// TIA Portal project "HEAT-1-CADIZ-V25" (V20) (continued)
VAR_GLOBAL   // PLC tag table "Robot Position"
   "tcpPosIniX_00" AT %I632.0 : Bool;   // $OUT[257]
   "tcpPosIniX_01" AT %I632.1 : Bool;
   "tcpPosIniX_02" AT %I632.2 : Bool;
   "tcpPosIniX_03" AT %I632.3 : Bool;
   "tcpPosIniX_04" AT %I632.4 : Bool;
   "tcpPosIniX_05" AT %I632.5 : Bool;
   "tcpPosIniX_06" AT %I632.6 : Bool;
   "tcpPosIniX_07" AT %I632.7 : Bool;
   "tcpPosIniX_08" AT %I633.0 : Bool;
   "tcpPosIniX_09" AT %I633.1 : Bool;
   "tcpPosIniX_10" AT %I633.2 : Bool;
   "tcpPosIniX_11" AT %I633.3 : Bool;
   "tcpPosIniX_12" AT %I633.4 : Bool;
   "tcpPosIniX_13" AT %I633.5 : Bool;
   "tcpPosIniX_14" AT %I633.6 : Bool;
   "tcpPosIniX_15" AT %I633.7 : Bool;
   "tcpPosIniX_16" AT %I634.0 : Bool;
   "tcpPosIniX_17" AT %I634.1 : Bool;
   "tcpPosIniX_18" AT %I634.2 : Bool;
   "tcpPosIniX_19" AT %I634.3 : Bool;
   "tcpPosIniX_20" AT %I634.4 : Bool;
   "tcpPosIniX_21" AT %I634.5 : Bool;
   "tcpPosIniX_22" AT %I634.6 : Bool;
   "tcpPosIniX_23" AT %I634.7 : Bool;
   "tcpPosIniX_24" AT %I635.0 : Bool;
   "tcpPosIniX_25" AT %I635.1 : Bool;
   "tcpPosIniX_26" AT %I635.2 : Bool;
   "tcpPosIniX_27" AT %I635.3 : Bool;
   "tcpPosIniX_28" AT %I635.4 : Bool;
   "tcpPosIniX_29" AT %I635.5 : Bool;
   "tcpPosIniX_30" AT %I635.6 : Bool;
   "tcpPosIniX_31" AT %I635.7 : Bool;
   "tcpPosIniY_00" AT %I636.0 : Bool;
   "tcpPosIniY_01" AT %I636.1 : Bool;
   "tcpPosIniY_02" AT %I636.2 : Bool;
   "tcpPosIniY_03" AT %I636.3 : Bool;
   "tcpPosIniY_04" AT %I636.4 : Bool;
   "tcpPosIniY_05" AT %I636.5 : Bool;
   "tcpPosIniY_06" AT %I636.6 : Bool;
   "tcpPosIniY_07" AT %I636.7 : Bool;
   "tcpPosIniY_08" AT %I637.0 : Bool;
   "tcpPosIniY_09" AT %I637.1 : Bool;
   "tcpPosIniY_10" AT %I637.2 : Bool;
   "tcpPosIniY_11" AT %I637.3 : Bool;
   "tcpPosIniY_12" AT %I637.4 : Bool;
   "tcpPosIniY_13" AT %I637.5 : Bool;
   "tcpPosIniY_14" AT %I637.6 : Bool;
   "tcpPosIniY_15" AT %I637.7 : Bool;
   "tcpPosIniY_16" AT %I638.0 : Bool;
   "tcpPosIniY_17" AT %I638.1 : Bool;
   "tcpPosIniY_18" AT %I638.2 : Bool;
   "tcpPosIniY_19" AT %I638.3 : Bool;
   "tcpPosIniY_20" AT %I638.4 : Bool;
   "tcpPosIniY_21" AT %I638.5 : Bool;
   "tcpPosIniY_22" AT %I638.6 : Bool;
   "tcpPosIniY_23" AT %I638.7 : Bool;
   "tcpPosIniY_24" AT %I639.0 : Bool;
   "tcpPosIniY_25" AT %I639.1 : Bool;
   "tcpPosIniY_26" AT %I639.2 : Bool;
   "tcpPosIniY_27" AT %I639.3 : Bool;
   "tcpPosIniY_28" AT %I639.4 : Bool;
   "tcpPosIniY_29" AT %I639.5 : Bool;
   "tcpPosIniY_30" AT %I639.6 : Bool;
   "tcpPosIniY_31" AT %I639.7 : Bool;
   "tcpPosIniZ_00" AT %I640.0 : Bool;
   "tcpPosIniZ_01" AT %I640.1 : Bool;
   "tcpPosIniZ_02" AT %I640.2 : Bool;
   "tcpPosIniZ_03" AT %I640.3 : Bool;
   "tcpPosIniZ_04" AT %I640.4 : Bool;
   "tcpPosIniZ_05" AT %I640.5 : Bool;
   "tcpPosIniZ_06" AT %I640.6 : Bool;
   "tcpPosIniZ_07" AT %I640.7 : Bool;
   "tcpPosIniZ_08" AT %I641.0 : Bool;
   "tcpPosIniZ_09" AT %I641.1 : Bool;
   "tcpPosIniZ_10" AT %I641.2 : Bool;
   "tcpPosIniZ_11" AT %I641.3 : Bool;
   "tcpPosIniZ_12" AT %I641.4 : Bool;
   "tcpPosIniZ_13" AT %I641.5 : Bool;
   "tcpPosIniZ_14" AT %I641.6 : Bool;
   "tcpPosIniZ_15" AT %I641.7 : Bool;
   "tcpPosIniZ_16" AT %I642.0 : Bool;
   "tcpPosIniZ_17" AT %I642.1 : Bool;
   "tcpPosIniZ_18" AT %I642.2 : Bool;
   "tcpPosIniZ_19" AT %I642.3 : Bool;
   "tcpPosIniZ_20" AT %I642.4 : Bool;
   "tcpPosIniZ_21" AT %I642.5 : Bool;
   "tcpPosIniZ_22" AT %I642.6 : Bool;
   "tcpPosIniZ_23" AT %I642.7 : Bool;
   "tcpPosIniZ_24" AT %I643.0 : Bool;
   "tcpPosIniZ_25" AT %I643.1 : Bool;
   "tcpPosIniZ_26" AT %I643.2 : Bool;
   "tcpPosIniZ_27" AT %I643.3 : Bool;
   "tcpPosIniZ_28" AT %I643.4 : Bool;
   "tcpPosIniZ_29" AT %I643.5 : Bool;
   "tcpPosIniZ_30" AT %I643.6 : Bool;
   "tcpPosIniZ_31" AT %I643.7 : Bool;
   "e1PosIni_00" AT %I644.0 : Bool;
   "e1PosIni_01" AT %I644.1 : Bool;
   "e1PosIni_02" AT %I644.2 : Bool;
   "e1PosIni_03" AT %I644.3 : Bool;
   "e1PosIni_04" AT %I644.4 : Bool;
   "e1PosIni_05" AT %I644.5 : Bool;
   "e1PosIni_06" AT %I644.6 : Bool;
   "e1PosIni_07" AT %I644.7 : Bool;
   "e1PosIni_08" AT %I645.0 : Bool;
   "e1PosIni_09" AT %I645.1 : Bool;
   "e1PosIni_10" AT %I645.2 : Bool;
   "e1PosIni_11" AT %I645.3 : Bool;
   "e1PosIni_12" AT %I645.4 : Bool;
   "e1PosIni_13" AT %I645.5 : Bool;
   "e1PosIni_14" AT %I645.6 : Bool;
   "e1PosIni_15" AT %I645.7 : Bool;
   "e1PosIni_16" AT %I646.0 : Bool;
   "e1PosIni_17" AT %I646.1 : Bool;
   "e1PosIni_18" AT %I646.2 : Bool;
   "e1PosIni_19" AT %I646.3 : Bool;
   "e1PosIni_20" AT %I646.4 : Bool;
   "e1PosIni_21" AT %I646.5 : Bool;
   "e1PosIni_22" AT %I646.6 : Bool;
   "e1PosIni_23" AT %I646.7 : Bool;
   "e1PosIni_24" AT %I647.0 : Bool;
   "e1PosIni_25" AT %I647.1 : Bool;
   "e1PosIni_26" AT %I647.2 : Bool;
   "e1PosIni_27" AT %I647.3 : Bool;
   "e1PosIni_28" AT %I647.4 : Bool;
   "e1PosIni_29" AT %I647.5 : Bool;
   "e1PosIni_30" AT %I647.6 : Bool;
   "e1PosIni_31" AT %I647.7 : Bool;
   "tcpPosFinX_00" AT %I648.0 : Bool;
   "tcpPosFinX_01" AT %I648.1 : Bool;
   "tcpPosFinX_02" AT %I648.2 : Bool;
   "tcpPosFinX_03" AT %I648.3 : Bool;
   "tcpPosFinX_04" AT %I648.4 : Bool;
   "tcpPosFinX_05" AT %I648.5 : Bool;
   "tcpPosFinX_06" AT %I648.6 : Bool;
   "tcpPosFinX_07" AT %I648.7 : Bool;
   "tcpPosFinX_08" AT %I649.0 : Bool;
   "tcpPosFinX_09" AT %I649.1 : Bool;
   "tcpPosFinX_10" AT %I649.2 : Bool;
   "tcpPosFinX_11" AT %I649.3 : Bool;
   "tcpPosFinX_12" AT %I649.4 : Bool;
   "tcpPosFinX_13" AT %I649.5 : Bool;
   "tcpPosFinX_14" AT %I649.6 : Bool;
   "tcpPosFinX_15" AT %I649.7 : Bool;
   "tcpPosFinX_16" AT %I650.0 : Bool;
   "tcpPosFinX_17" AT %I650.1 : Bool;
   "tcpPosFinX_18" AT %I650.2 : Bool;
   "tcpPosFinX_19" AT %I650.3 : Bool;
   "tcpPosFinX_20" AT %I650.4 : Bool;
   "tcpPosFinX_21" AT %I650.5 : Bool;
   "tcpPosFinX_22" AT %I650.6 : Bool;
   "tcpPosFinX_23" AT %I650.7 : Bool;
   "tcpPosFinX_24" AT %I651.0 : Bool;
   "tcpPosFinX_25" AT %I651.1 : Bool;
   "tcpPosFinX_26" AT %I651.2 : Bool;
   "tcpPosFinX_27" AT %I651.3 : Bool;
   "tcpPosFinX_28" AT %I651.4 : Bool;
   "tcpPosFinX_29" AT %I651.5 : Bool;
   "tcpPosFinX_30" AT %I651.6 : Bool;
   "tcpPosFinX_31" AT %I651.7 : Bool;
   "tcpPosFinY_00" AT %I652.0 : Bool;
   "tcpPosFinY_01" AT %I652.1 : Bool;
   "tcpPosFinY_02" AT %I652.2 : Bool;
   "tcpPosFinY_03" AT %I652.3 : Bool;
   "tcpPosFinY_04" AT %I652.4 : Bool;
   "tcpPosFinY_05" AT %I652.5 : Bool;
   "tcpPosFinY_06" AT %I652.6 : Bool;
   "tcpPosFinY_07" AT %I652.7 : Bool;
   "tcpPosFinY_08" AT %I653.0 : Bool;
   "tcpPosFinY_09" AT %I653.1 : Bool;
   "tcpPosFinY_10" AT %I653.2 : Bool;
   "tcpPosFinY_11" AT %I653.3 : Bool;
   "tcpPosFinY_12" AT %I653.4 : Bool;
   "tcpPosFinY_13" AT %I653.5 : Bool;
   "tcpPosFinY_14" AT %I653.6 : Bool;
   "tcpPosFinY_15" AT %I653.7 : Bool;
   "tcpPosFinY_16" AT %I654.0 : Bool;
   "tcpPosFinY_17" AT %I654.1 : Bool;
   "tcpPosFinY_18" AT %I654.2 : Bool;
   "tcpPosFinY_19" AT %I654.3 : Bool;
   "tcpPosFinY_20" AT %I654.4 : Bool;
   "tcpPosFinY_21" AT %I654.5 : Bool;
   "tcpPosFinY_22" AT %I654.6 : Bool;
   "tcpPosFinY_23" AT %I654.7 : Bool;
   "tcpPosFinY_24" AT %I655.0 : Bool;
   "tcpPosFinY_25" AT %I655.1 : Bool;
   "tcpPosFinY_26" AT %I655.2 : Bool;
   "tcpPosFinY_27" AT %I655.3 : Bool;
   "tcpPosFinY_28" AT %I655.4 : Bool;
   "tcpPosFinY_29" AT %I655.5 : Bool;
   "tcpPosFinY_30" AT %I655.6 : Bool;
   "tcpPosFinY_31" AT %I655.7 : Bool;
   "tcpPosE1_01" AT %I628.0 : Bool;
   "tcpPosE1_02" AT %I628.1 : Bool;
   "tcpPosE1_03" AT %I628.2 : Bool;
   "tcpPosE1_04" AT %I628.3 : Bool;
   "tcpPosE1_05" AT %I628.4 : Bool;
   "tcpPosE1_06" AT %I628.5 : Bool;
   "tcpPosE1_07" AT %I628.6 : Bool;
   "tcpPosE1_08" AT %I628.7 : Bool;
   "tcpPosE1_09" AT %I629.0 : Bool;
   "tcpPosE1_10" AT %I629.1 : Bool;
   "tcpPosE1_11" AT %I629.2 : Bool;
   "tcpPosE1_12" AT %I629.3 : Bool;
   "tcpPosE1_13" AT %I629.4 : Bool;
   "tcpPosE1_14" AT %I629.5 : Bool;
   "tcpPosE1_15" AT %I629.6 : Bool;
   "tcpPosE1_16" AT %I629.7 : Bool;
   "tcpPosE1_17" AT %I630.0 : Bool;
   "tcpPosE1_18" AT %I630.1 : Bool;
   "tcpPosE1_19" AT %I630.2 : Bool;
   "tcpPosE1_20" AT %I630.3 : Bool;
   "tcpPosE1_21" AT %I630.4 : Bool;
   "tcpPosE1_22" AT %I630.5 : Bool;
   "tcpPosE1_23" AT %I630.6 : Bool;
   "tcpPosE1_24" AT %I630.7 : Bool;
   "tcpPosE1_25" AT %I631.0 : Bool;
   "tcpPosE1_26" AT %I631.1 : Bool;
   "tcpPosE1_27" AT %I631.2 : Bool;
   "tcpPosE1_28" AT %I631.3 : Bool;
   "tcpPosE1_29" AT %I631.4 : Bool;
   "tcpPosE1_30" AT %I631.5 : Bool;
   "tcpPosE1_31" AT %I631.6 : Bool;
   "tcpPosE1_32" AT %I631.7 : Bool;
   "tcpPosIniX_rawLe32" AT %ID632 : DWord;
   "tcpPosIniY_rawLe32" AT %ID636 : DWord;
   "tcpPosIniZ_rawLe32" AT %ID640 : DWord;
   "tcpPosFinX_rawLe32" AT %ID648 : DWord;
   "tcpPosFinY_rawLe32" AT %ID652 : DWord;
   "e1_rawLe32" AT %ID628 : DWord;
   "e1PosIni_rawLe32" AT %ID644 : DWord;
   "tcpPosFinZ_rawLe32" AT %ID656 : DWord;
   "e1PosFin_rawLe32" AT %ID660 : DWord;
END_VAR

VAR_GLOBAL   // PLC tag table "Tool Change"
   "dockSensorToolYugoInPosition" AT %I150.0 : Bool;   // DETECTOR_YUGO_LP
   "dockSensorCoverYugoClosed" AT %I150.1 : Bool;   // TAPA_CERRADA_YUGO_LP
   "dockSensorCoverOpen" AT %I160.0 : Bool;   // TAPA_ABIERTA_YUGO_LP
   "dockValveV2UnlockOnYugo" AT %Q171.2 : Bool;   // SOLTAR_HERRAMIENTA_YUGO_LP / CAMBIA A FALSE
   "dockValveCoverOpenOn" AT %Q170.0 : Bool;   // ABRIR_TAPA_YUGO_LP
   "dockValveCoverCloseOn" AT %Q170.1 : Bool;   // CERRAR_TAPA_YUGO_LP
   "robotSensorMpsUnlocked" AT %I200.0 : Bool;   // INTERCAMBIO_DESBLOQUEADO_LR
   "robotSensorMpsLocked" AT %I200.1 : Bool;   // INTERCAMBIO_BLOQUEADO_LR
   "robotSensorMpsCoupled" AT %I200.2 : Bool;   // HERRAMIENTA_PUESTA_LR /AL COLOCAR METAL
   "robotSensorMpsCtrlAirPressureOk" AT %I200.3 : Bool;   // PRESION_CORRECTA_LR
   "toolReqId_01" AT %Q618.1 : Bool;   // INKUKA_DETECTOR_HERRAMIENTA
   "toolReqId_02" AT %Q618.2 : Bool;   // INKUKA_TAPA_CERRADA_YUGO
   "toolReqId_03" AT %Q618.3 : Bool;   // INKUKA_TAPA_ABIERTA_YUGO
   "toolReqId_04" AT %Q618.4 : Bool;   // INKUKA_INTERCAMBIO_DESBLOQUEADO
   "toolReqId_05" AT %Q618.5 : Bool;   // INKUKA_INTERCAMBIO_BLOQUEADO
   "toolReqId_06" AT %Q618.6 : Bool;   // INKUKA_HERRAMIENTA_PUESTA /AL COLOCAR util met
   "toolReqId_07" AT %Q618.7 : Bool;
   "kukaCmdUnlockMpsYugo" AT %I696.0 : Bool;   // OUTKUKA_SOLTAR_HERRAMIENTA_YUGO
   "kukaCmdOpenCover" AT %I696.1 : Bool;   // OUTKUKA_ABRIR_TAPA_YUGO
   "kukaCmdCloseCover" AT %I696.2 : Bool;   // OUTKUKA_CERRAR_TAPA_YUGO
   "V1_B14_S2" AT %Q0.0 : Bool;   // Anticolision - OPR
   "V1_B12_S4" AT %Q0.1 : Bool;   // Mps Bloqueo SIL 2
   "V2_B14_S2" AT %Q0.2 : Bool;
   "V2_B12_S4" AT %Q0.3 : Bool;
   "toolReqId_00" AT %Q618.0 : Bool;
   "toolReqId_08" AT %Q619.0 : Bool;
   "toolReqId_09" AT %Q619.1 : Bool;
   "toolReqId_10" AT %Q619.2 : Bool;
   "toolReqId_11" AT %Q619.3 : Bool;
   "toolReqId_12" AT %Q619.4 : Bool;
   "toolReqId_13" AT %Q619.5 : Bool;
   "toolReqId_14" AT %Q619.6 : Bool;
   "toolReqId_15" AT %Q619.7 : Bool;
   "toolReqId" AT %QW618 : Word;
   "baseReqId" AT %QW620 : Word;
   "kukaFeedbackDockToolYugoInPosition" AT %Q696.4 : Bool;   // $IN[773]
   "kukaFeedbackDockYugoCoverClosed" AT %Q696.5 : Bool;
   "kukaFeedbackDockYugoCoverOpen" AT %Q696.6 : Bool;
   "kukaFeedbackRobotMpsUnlocked" AT %Q696.0 : Bool;   // $IN[769]
   "kukaFeedbackRobotMpsLocked" AT %Q696.1 : Bool;
   "kukaFeedbackRobotMpsCoupled" AT %Q696.2 : Bool;
   "kukaFeedbackRobotMpsCtrlAirPressureOk" AT %Q696.3 : Bool;
   "dockValveV2UnlockOnPepa" AT %Q171.4 : Bool;   // SOLTAR_HERRAMIENTA_PEPA
   "dockSensorToolPepaInPosition" AT %I150.2 : Bool;
   "kukaCmdSafeForChange" AT %I696.3 : Bool;   // $OUT[772]
   "kukaCmdUnlockMpsPepa" AT %I696.4 : Bool;   // $OUT[773]
   "kukaCmdOpenCoverPepa" AT %I696.5 : Bool;   // $OUT[774]
   "kukaCmdUnlockMpsMarker" AT %I696.7 : Bool;   // $OUT[775]
   "kukaCmdOpenCoverMarker" AT %I697.0 : Bool;   // $OUT[776]
   "kukaCmdCloseCoverMarker" AT %I697.1 : Bool;   // $OUT[777]
   "kukaCmdUnlockMpsGocator" AT %I697.2 : Bool;
   "kukaCmdOpenCoverGocator" AT %I697.3 : Bool;
   "kukaCmdCloseCoverGocator" AT %I697.4 : Bool;
   "kukaCmdCloseCoverPepa" AT %I696.6 : Bool;
   "kukaCmdUnlockMpsPole" AT %I697.5 : Bool;
   "kukaCmdOpenCoverPole" AT %I697.6 : Bool;
   "kukaCmdCloseCoverPole" AT %I697.7 : Bool;
   "kukaFeedbackDockToolPepaInPosition" AT %Q696.7 : Bool;
   "kukaFeedbackDockPepaCoverClosed" AT %Q697.0 : Bool;
   "kukaFeedbackDockPepaCoverOpen" AT %Q697.1 : Bool;
   "kukaFeedbackDockToolMarkerInPosition" AT %Q697.2 : Bool;
   "kukaFeedbackDockMarkerCoverClosed" AT %Q697.3 : Bool;
   "kukaFeedbackDockMarkerCoverOpen" AT %Q697.4 : Bool;
   "kukaFeedbackDockToolGocatorInPosition" AT %Q697.5 : Bool;
   "kukaFeedbackDockGocatorCoverClosed" AT %Q697.6 : Bool;
   "kukaFeedbackDockGocatorCoverOpen" AT %Q697.7 : Bool;
   "kukaFeedbackDockToolPoleInPosition" AT %Q698.0 : Bool;
   "kukaFeedbackDockPoleCoverClosed" AT %Q698.1 : Bool;
   "kukaFeedbackDockPoleCoverOpen" AT %Q698.2 : Bool;
   "dockSensorCoverPepaClosed" AT %I150.3 : Bool;
   "dockSensorToolPoleInPosition" AT %I150.4 : Bool;
   "dockSensorToolMarkerInPosition" AT %I150.6 : Bool;
   "dockSensorToolGocatorInPosition" AT %I151.0 : Bool;
   "pruebaHerramienta2enStand" AT %I151.2 : Bool;
   "pruebaHerramienta1enStand" AT %I151.1 : Bool;
   "pruebaHerramienta3enStand" AT %I151.3 : Bool;
   "pruebaHerramienta4enStand" AT %I151.4 : Bool;
   "pruebaHerramient54enStand" AT %I150.7 : Bool;
   "dockSensorTooPole%I150.5InPosition" AT %I150.5 : Bool;
END_VAR

VAR_GLOBAL   // PLC tag table "General"
   "ALM_PRESS_SENSOR" AT %I10.0 : Bool;   // Pressure-sensor alarm
   "CMD_TANK_FILL" AT %Q30.0 : Bool;   // LLENAR CUBA
   "CMD_TANK_DRAIN" AT %Q30.1 : Bool;   // VACIAR CUBA
   "RECIRCULACION" AT %Q30.2 : Bool;   // CONMUTADOR MANUAL / cambiado a recirculacion
END_VAR

VAR_GLOBAL   // PLC tag table "Tag table_1"
   "Sensor_plato_giro_1" AT %I410.0 : Bool;
   "Sensor_Plato_giro_2" AT %I410.1 : Bool;
   "Sensor_plato_giro_3" AT %I410.2 : Bool;
   "Sensor_ADN_bastidor_bloqueado_1" AT %I410.3 : Bool;
   "Sensor_ADN_bastidor_desbloqueado_1" AT %I410.4 : Bool;
   "Sensor_ADN_bastidor_bloqueado_2" AT %I410.5 : Bool;
   "Sensor_ADN_bastidor_desbloqueado_2" AT %I410.6 : Bool;
   "SENSOR_CRDSNU_BASTIDOR_BLOQUEADO_1" AT %I410.7 : Bool;
   "SENSOR_CRDSNU_BASTIDOR_DESBLOQUEADO_1" AT %I411.0 : Bool;
   "SENSOR_CRDSNU_BASTIDOR_BLOQUEADO_2" AT %I411.1 : Bool;
   "SENSOR_CRDSNU_BASTIDOR_DESBLOQUEADO_2" AT %I411.2 : Bool;
   "SENSOR_DSBG_BASTIDOR_ARRIBA_1" AT %I411.3 : Bool;
   "SENSOR_DSBG_BASTIDOR_ABAJO_1" AT %I411.4 : Bool;
   "SENSOR_DSBG_BASTIDOR_ARRIBA_2" AT %I411.5 : Bool;
   "SENSOR_DSBG_BASTIDOR_ABAJO_2" AT %I411.6 : Bool;
   "PULSADOR_SUBIR_1" AT %I412.0 : Bool;
   "PULSADOR_BAJAR_1" AT %I412.1 : Bool;
   "PULSADOR_SUBIR_2" AT %I412.2 : Bool;
   "PULSADOR_BAJAR_2" AT %I412.3 : Bool;
   "VALVULA_52_BIESTABLE_11" AT %Q420.0 : Bool;
   "VALVULA_52_BIESTABLE_12" AT %Q420.1 : Bool;
   "VALVULA_52_BIESTABLE_21" AT %Q420.2 : Bool;
   "VALVULA_52_BIESTABLE_22" AT %Q420.3 : Bool;
   "VÁLVULA_52_MONOESTABLE_1" AT %Q420.4 : Bool;
   "VÁLVULA_52_MONOESTABLE_2" AT %Q420.5 : Bool;
   "VÁLVULA_52_MONOESTABLE_3" AT %Q420.6 : Bool;
   "VÁLVULA_52_MONOESTABLE_4" AT %Q420.7 : Bool;
   "VÁLVULA_52_MONOESTABLE_5" AT %Q421.0 : Bool;
   "SENSOR_DSBG_BASTIDOR_ABAJO_3" AT %I411.7 : Bool;
   "PULSADOR_BAJAR_3" AT %I412.4 : Bool;
   "PULSADOR_BAJAR_4" AT %I412.5 : Bool;
   "PULSADOR_BAJAR_5" AT %I412.6 : Bool;
   "PULSADOR_BAJAR_6" AT %I412.7 : Bool;
   "PULSADOR_BAJAR_7" AT %I413.0 : Bool;
   "PULSADOR_BAJAR_8" AT %I413.1 : Bool;
   "PULSADOR_BAJAR_9" AT %I413.2 : Bool;
   "PULSADOR_BAJAR_10" AT %I413.3 : Bool;
   "PULSADOR_BAJAR_11" AT %I413.4 : Bool;
   "PULSADOR_BAJAR_12" AT %I413.5 : Bool;
   "PULSADOR_BAJAR_13" AT %I413.6 : Bool;
   "PULSADOR_BAJAR_14" AT %I413.7 : Bool;
   "VÁLVULA_52_MONOESTABLE_6" AT %Q421.1 : Bool;
   "VÁLVULA_52_MONOESTABLE_7" AT %Q421.2 : Bool;
   "VÁLVULA_52_MONOESTABLE_8" AT %Q421.3 : Bool;
   "VÁLVULA_52_MONOESTABLE_9" AT %Q421.4 : Bool;
   "VÁLVULA_52_MONOESTABLE_10" AT %Q421.5 : Bool;
   "VÁLVULA_52_MONOESTABLE_11" AT %Q421.6 : Bool;
   "VÁLVULA_52_MONOESTABLE_12" AT %Q421.7 : Bool;
   "VÁLVULA_52_MONOESTABLE_13" AT %Q422.0 : Bool;
   "VÁLVULA_52_MONOESTABLE_14" AT %Q422.1 : Bool;
   "VÁLVULA_52_MONOESTABLE_15" AT %Q422.2 : Bool;
   "VÁLVULA_52_MONOESTABLE_16" AT %Q422.3 : Bool;
   "VÁLVULA_52_MONOESTABLE_17" AT %Q422.4 : Bool;
   "VÁLVULA_52_MONOESTABLE_18" AT %Q422.5 : Bool;
   "VÁLVULA_52_MONOESTABLE_19" AT %Q422.6 : Bool;
   "VÁLVULA_52_MONOESTABLE_20" AT %Q422.7 : Bool;
   "VÁLVULA_52_MONOESTABLE_21" AT %Q423.0 : Bool;
   "VÁLVULA_52_MONOESTABLE_22" AT %Q423.1 : Bool;
   "VÁLVULA_52_MONOESTABLE_23" AT %Q423.2 : Bool;
   "VÁLVULA_52_MONOESTABLE_24" AT %Q423.3 : Bool;
   "VÁLVULA_52_MONOESTABLE_25" AT %Q423.4 : Bool;
   "VÁLVULA_52_MONOESTABLE_26" AT %Q423.5 : Bool;
   "VÁLVULA_52_MONOESTABLE_27" AT %Q423.6 : Bool;
   "VÁLVULA_52_MONOESTABLE_28" AT %Q423.7 : Bool;
END_VAR

TYPE "UDT_Dock"
   STRUCT
      Sensor : Struct
         CoverOpen : Bool;
         CoverClosed : Bool;
         ToolInPosition : Bool;
      END_STRUCT;
      Valve : Struct
         CoverOpenOn : Bool;
         CoverCloseOn : Bool;
         V2UnlockOn : Bool;
      END_STRUCT;
   END_STRUCT;
END_TYPE

TYPE "UDT_RobotMps"
   STRUCT
      Sensor : Struct
         Coupled : Bool;
         Locked : Bool;
         Unlocked : Bool;
         CtrlAirPressureOk : Bool;
      END_STRUCT;
   END_STRUCT;
END_TYPE

// folder: 10. System

DATA_BLOCK "HMI_CUBA_DB"   // DB17
{ S7_Optimized_Access := 'TRUE' }
VERSION : 0.1
// stored: InstanceOfName HMI_CUBA
"HMI_CUBA"
BEGIN
END_DATA_BLOCK

DATA_BLOCK "instKukaControlSeq_DB"   // DB20
{ S7_Optimized_Access := 'TRUE' }
VERSION : 0.1
// stored: InstanceOfName KukaControlSeq
"KukaControlSeq"
BEGIN
END_DATA_BLOCK

DATA_BLOCK "GIRO_POSITIVO_DB"   // DB27
{ S7_Optimized_Access := 'TRUE' }
VERSION : 0.1
// stored: InstanceOfName GIRO_POSITIVO
"GIRO_POSITIVO"
BEGIN
END_DATA_BLOCK

DATA_BLOCK "GIRO_NEGATIVO_1_DB"   // DB28
{ S7_Optimized_Access := 'TRUE' }
VERSION : 0.1
// stored: InstanceOfName GIRO_NEGATIVO_1
"GIRO_NEGATIVO_1"
BEGIN
END_DATA_BLOCK

// folder: 10. System/DbsInstancia

DATA_BLOCK "InstKukaControlSeq"   // DB14
{ S7_Optimized_Access := 'TRUE' }
VERSION : 0.1
// stored: InstanceOfName KukaControlSeq
"KukaControlSeq"
BEGIN
END_DATA_BLOCK

DATA_BLOCK "InstSupervisorSeq"   // DB15
{ S7_Optimized_Access := 'TRUE' }
VERSION : 0.1
// stored: InstanceOfName SupervisorSeq
"SupervisorSeq"
BEGIN
END_DATA_BLOCK

DATA_BLOCK "InstSeqManager"   // DB16
{ S7_Optimized_Access := 'TRUE' }
VERSION : 0.1
// stored: InstanceOfName SeqManager
"SeqManager"
BEGIN
END_DATA_BLOCK

DATA_BLOCK "AutoExtSeq_DB"   // DB18
{ S7_Optimized_Access := 'TRUE' }
VERSION : 0.1
// stored: InstanceOfName AutoExtSeq
"AutoExtSeq"
BEGIN
END_DATA_BLOCK

DATA_BLOCK "instSupervisorSeq_DB"   // DB21
{ S7_Optimized_Access := 'TRUE' }
VERSION : 0.1
// stored: InstanceOfName SupervisorSeq
"SupervisorSeq"
BEGIN
END_DATA_BLOCK

// folder: 10. System/DbsOpcUa

DATA_BLOCK "PlcStatus"   // DB4
{ S7_Optimized_Access := 'TRUE' }
VERSION : 0.1
   VAR
      "- FOR  KUKACONTROL-" : Bool;
      mode : Struct
         effective : UInt;
         ready : Bool;
      END_STRUCT;
      active : Struct
         baseId : UInt;
         toolId : UInt;
         profileId : UInt;
      END_STRUCT;
      exec : Struct
         ackSeq : UInt;
         accepted : Bool;
         busy : Bool;
         done : Bool;
         error : Bool;
         errorCode : UDInt;
         cancelAck : Bool;
         pauseAck : Bool;
         resumeAck : Bool;
         paused : Bool;
      END_STRUCT;
      pose : Struct
         tcpPosX_mm : LReal;
         tcpPosY_mm : LReal;
         tcpPosZ_mm : LReal;
         tcpOriA_deg : LReal;
         tcpOriB_deg : LReal;
         tcpOriC_deg : LReal;
         e1Pos_mm : LReal;
      END_STRUCT;
      teach : Struct
         startX_mm : LReal;
         startY_mm : LReal;
         startZ_mm : LReal;
         startE1_mm : LReal;
         startOk : Bool;
         endX_mm : LReal;
         endY_mm : LReal;
         endZ_mm : LReal;
         endE1_mm : LReal;
         endOk : Bool;
      END_STRUCT;
      systemArmed : Bool;
      robotInHome : Bool;
      robotInAutExt : Bool;
      heartbeatPlc : Bool;
      stepPlc : Int;
      plcOk : Bool := true;
      safetyOk : Bool := true;
      airOk : Bool := true;
      inspWaterOk : Bool := true;
      tankWaterOk : Bool := true;
      robotOk : Bool := true;
      acknowledge : Bool;
      carriageId : String;
      newCarriageId : Bool;
      idRunning : Bool;
      idOk : Bool;
      startUsReady : Bool;
      stopUsReady : Bool;
      paCheckReady : Bool;
      gainReady : Bool;
      tcgReady : Bool;
      idScan : String;
      pointOrigin : LReal;
      xSize : LReal;
      ySize : LReal;
      scanRefStart : Bool;
      scanInspStart : Bool;
      markRunning : Bool;
      markState : Bool;
      breakUs : Bool;
      unbreakUs : Bool;
      robotRescanning : Bool;
      acknowledgeError : Bool;
   END_VAR
BEGIN
END_DATA_BLOCK

DATA_BLOCK "KukaControlCmd"   // DB5
{ S7_Optimized_Access := 'TRUE' }
VERSION : 0.1
   VAR
      code : UInt;
      seq : UInt;
      tcpTargetX_mm : LReal;
      tcpTargetY_mm : LReal;
      tcpTargetZ_mm : LReal;
      e1Target : LReal;
      toolRequestId : UInt;
      baseRequestId : UInt;
      profileRequestId : UInt;
      vel_mms : UInt;
      index_mm : UInt;
      apo_mm : LReal;
      programRequestId : UInt;
      cancelGo : Bool;
      pauseGo : Bool;
      resumeGo : Bool;
      mode : Struct
         request : UInt;
         reqSeq : UInt;
      END_STRUCT;
      scanPuntoInicialX : LReal;
      scanPuntoInicialY : LReal;
      scanPuntoInicialZ : LReal;
      scanPuntoInicialE1 : LReal;
      scanPuntoFinalX : LReal;
      scanPuntoFinalY : LReal;
      scanPuntoFinalZ : LReal;
      scanPuntoFinalE1 : LReal;
      carriageId : String;
      qrReady : Bool;
   END_VAR
BEGIN
END_DATA_BLOCK

DATA_BLOCK "SupervisorCmd"   // DB6
{ S7_Optimized_Access := 'TRUE' }
VERSION : 0.1
   VAR
      heartbeatSupervisor : Bool;
      stepSupervisor : Int;
      supervisorOk : Bool := true;
      stateUs : Bool;
      reqCarriageId : Bool;
      reqId : Bool;
      pns : String;
      referencePart : String;
      endEffector : Int;
      utTech : UInt;
      teachReq : Bool;
      paCheckReq : Bool;
      tcgReq : Bool;
      startUsRunning : Bool;
      stopUsRunning : Bool;
      elemState : Bool;
      elemRunning : Bool;
      balState : Bool;
      balRunning : Bool;
      gainState : Bool;
      gainRunning : Bool;
      tcgInProgress : Bool;
      tcgNextStep : Bool;
      tcgState : Bool;
      reqRefPart : Bool;
      reqStopCycle : Bool;
      reqTcgAdj : Bool;
      scanRefState : Bool;
      scanRefRunning : Bool;
      reqPreEval : Bool;
      reqIdentificationState : Bool;
      scanInspState : Bool;
      scanInsprunning : Bool;
      reqMark : Bool;
      reqVerif : Bool;
      pointCoordinates : LReal;
      goBack : Bool;
      rescanning : Bool;
      errorMessage : String;
      errorOcurred : Bool;
      gainAdjustmentReq : Bool;
   END_VAR
BEGIN
END_DATA_BLOCK

// folder: 10. System/Utilities

DATA_BLOCK "Utilidades"   // DB37
{ S7_Optimized_Access := 'TRUE' }
VERSION : 0.1
   VAR
      numProg : USInt;
   END_VAR
BEGIN
END_DATA_BLOCK

// folder: 20. Robot Services/AutoExt

DATA_BLOCK "instAutoExtSeq"   // DB7
{ S7_Optimized_Access := 'TRUE' }
VERSION : 0.1
// stored: InstanceOfName AutoExtSeq
"AutoExtSeq"
BEGIN
END_DATA_BLOCK

// folder: 20. Robot Services/DbsInstancia

DATA_BLOCK "InstTcpJogging"   // DB2
{ S7_Optimized_Access := 'TRUE' }
VERSION : 0.1
// stored: InstanceOfName TcpJogging
"TcpJogging"
BEGIN
END_DATA_BLOCK

DATA_BLOCK "ToolChangeFork_DB"   // DB8
{ S7_Optimized_Access := 'TRUE' }
VERSION : 0.1
// stored: InstanceOfName ToolChange
"ToolChange"
BEGIN
END_DATA_BLOCK

DATA_BLOCK "TcpPoseDecoderLe32_DB"   // DB10
{ S7_Optimized_Access := 'TRUE' }
VERSION : 0.1
// stored: InstanceOfName TcpPoseDecoderLe32
"TcpPoseDecoderLe32"
BEGIN
END_DATA_BLOCK

DATA_BLOCK "InstTcpTarget"   // DB13
{ S7_Optimized_Access := 'TRUE' }
VERSION : 0.1
// stored: InstanceOfName TcpTarget
"TcpTarget"
BEGIN
END_DATA_BLOCK

// folder: 20. Robot Services/Tooling & Parking

DATA_BLOCK "ToolChangePepa"   // DB11
{ S7_Optimized_Access := 'TRUE' }
VERSION : 0.1
// stored: InstanceOfName ToolChange
"ToolChange"
BEGIN
END_DATA_BLOCK

DATA_BLOCK "MpsDockingStation_DB"   // DB22
{ S7_Optimized_Access := 'TRUE' }
VERSION : 0.1
// stored: InstanceOfName MpsDockingStation
"MpsDockingStation"
BEGIN
END_DATA_BLOCK

DATA_BLOCK "ToolChangePole_DB"   // DB23
{ S7_Optimized_Access := 'TRUE' }
VERSION : 0.1
// stored: InstanceOfName ToolChange
"ToolChange"
BEGIN
END_DATA_BLOCK

DATA_BLOCK "ToolInRobot_DB"   // DB32
{ S7_Optimized_Access := 'TRUE' }
VERSION : 0.1
// stored: InstanceOfName ToolInRobot
"ToolInRobot"
BEGIN
END_DATA_BLOCK

// folder: 30. Safety

DATA_BLOCK "InstMainSafety"   // DB1, F_DB
{ S7_Optimized_Access := 'TRUE' }
NAME : FUSI
VERSION : 0.1
// stored: InstanceOfName MainSafety
"MainSafety"
BEGIN
END_DATA_BLOCK

DATA_BLOCK "SafetyRobotDb"   // DB3, F_DB
{ S7_Optimized_Access := 'TRUE' }
VERSION : 0.1
BEGIN
END_DATA_BLOCK

// folder: 410. Festo cuba

DATA_BLOCK "HMI_CUBA_FESTO"   // DB12
{ S7_Optimized_Access := 'TRUE' }
VERSION : 0.1
   VAR
      HMI_Sensor_plato_giro_1 : Bool;
      HMI_Sensor_Plato_giro_2 : Bool;
      HMI_Sensor_plato_giro_3 : Bool;
      HMI_Sensor_ADN_bastidor_bloqueado_1 : Bool;
      HMI_Sensor_ADN_bastidor_desbloqueado_1 : Bool;
      HMI_Sensor_ADN_bastidor_bloqueado_2 : Bool;
      HMI_Sensor_ADN_bastidor_desbloqueado_2 : Bool;
      HMI_SENSOR_CRDSNU_BASTIDOR_BLOQUEADO_1 : Bool;
      HMI_SENSOR_CRDSNU_BASTIDOR_DESBLOQUEADO_1 : Bool;
      HMI_SENSOR_CRDSNU_BASTIDOR_BLOQUEADO_2 : Bool;
      HMI_SENSOR_CRDSNU_BASTIDOR_DESBLOQUEADO_2 : Bool;
      HMI_SENSOR_DSBG_BASTIDOR_ARRIBA_1 : Bool;
      HMI_SENSOR_DSBG_BASTIDOR_ABAJO_1 : Bool;
      HMI_SENSOR_DSBG_BASTIDOR_ARRIBA_2 : Bool;
      HMI_SENSOR_DSBG_BASTIDOR_ABAJO_2 : Bool;
      HMI_PULSADOR_SUBIR_1 : Bool;
      HMI_PULSADOR_BAJAR_1 : Bool;
      HMI_PULSADOR_SUBIR_2 : Bool;
      HMI_PULSADOR_BAJAR_2 : Bool;
      HMI_PULSADOR_BAJAR_3 : Bool;
      HMI_PULSADOR_BAJAR_4 : Bool;
      HMI_PULSADOR_BAJAR_5 : Bool;
      HMI_PULSADOR_BAJAR_6 : Bool;
      HMI_PULSADOR_BAJAR_7 : Bool;
      HMI_PULSADOR_BAJAR_8 : Bool;
      HMI_PULSADOR_BAJAR_9 : Bool;
      HMI_PULSADOR_BAJAR_10 : Bool;
      HMI_PULSADOR_BAJAR_11 : Bool;
      HMI_PULSADOR_BAJAR_12 : Bool;
      HMI_PULSADOR_BAJAR_13 : Bool;
      HMI_PULSADOR_BAJAR_14 : Bool;
      HMI_VALVULA_52_BIESTABLE_11 : Bool;
      HMI_VALVULA_52_BIESTABLE_12 : Bool;
      HMI_VALVULA_52_BIESTABLE_21 : Bool;
      HMI_VALVULA_52_BIESTABLE_22 : Bool;
      HMI_VÁLVULA_52_MONOESTABLE_1 : Bool;
      HMI_VÁLVULA_52_MONOESTABLE_2 : Bool;
      HMI_VÁLVULA_52_MONOESTABLE_3 : Bool;
      HMI_VÁLVULA_52_MONOESTABLE_4 : Bool;
      HMI_VÁLVULA_52_MONOESTABLE_5 : Bool;
      HMI_VÁLVULA_52_MONOESTABLE_6 : Bool;
      HMI_VÁLVULA_52_MONOESTABLE_7 : Bool;
      HMI_VÁLVULA_52_MONOESTABLE_8 : Bool;
      HMI_VÁLVULA_52_MONOESTABLE_9 : Bool;
      HMI_VÁLVULA_52_MONOESTABLE_10 : Bool;
      HMI_VÁLVULA_52_MONOESTABLE_11 : Bool;
      HMI_VÁLVULA_52_MONOESTABLE_12 : Bool;
      HMI_VÁLVULA_52_MONOESTABLE_13 : Bool;
      HMI_VÁLVULA_52_MONOESTABLE_14 : Bool;
      HMI_VÁLVULA_52_MONOESTABLE_15 : Bool;
      HMI_VÁLVULA_52_MONOESTABLE_16 : Bool;
      HMI_VÁLVULA_52_MONOESTABLE_17 : Bool;
      HMI_VÁLVULA_52_MONOESTABLE_18 : Bool;
      HMI_VÁLVULA_52_MONOESTABLE_19 : Bool;
      HMI_VÁLVULA_52_MONOESTABLE_20 : Bool;
      HMI_VÁLVULA_52_MONOESTABLE_21 : Bool;
      HMI_VÁLVULA_52_MONOESTABLE_22 : Bool;
      HMI_VÁLVULA_52_MONOESTABLE_23 : Bool;
      HMI_VÁLVULA_52_MONOESTABLE_24 : Bool;
      HMI_VÁLVULA_52_MONOESTABLE_25 : Bool;
      HMI_VÁLVULA_52_MONOESTABLE_26 : Bool;
      HMI_VÁLVULA_52_MONOESTABLE_27 : Bool;
      HMI_VÁLVULA_52_MONOESTABLE_28 : Bool;
      Estado_giro_pos_1 : Bool;
      Estado_giro_pos_2 : Bool;
      Estado_giro_pos_3 : Bool;
      Estado_giro_pos_4 : Bool;
      Estado_giro_neg_1 : Bool;
      Estado_giro_neg_2 : Bool;
      Estado_giro_neg_3 : Bool;
      Estado_giro_neg_4 : Bool;
      Estado_giro_neg_0 : Bool := true;
      Estado_giro_pos_0 : Bool := true;
      GIRO_AUTOMATICO_HABILITADO : Bool;
      Giro_negativo_auto : Bool;
      Giro_positivo_auto : Bool;
   END_VAR
BEGIN
END_DATA_BLOCK

// folder: Achim

DATA_BLOCK "Achim_testPepaFrk_DB"   // DB19
{ S7_Optimized_Access := 'TRUE' }
VERSION : 0.1
// stored: InstanceOfName Achim_testPepaFrk
"Achim_testPepaFrk"
BEGIN
END_DATA_BLOCK

// folder: Eliminar

DATA_BLOCK "DB_Supervisor"   // DB9
{ S7_Optimized_Access := 'TRUE' }
VERSION : 0.1
   VAR
      Common : Struct
         plc_ok : Bool;
         supervisor_ok : Bool;
         system_ok : Bool;
         safety_ok : Bool;
         air_ok : Bool;
         insp_water_ok : Bool;
         tank_water_ok : Bool;
         robot_ok : Bool;
         step_plc : Int;
         step_supervisor : Int;
         error : Bool;
         reset_req : Bool;
      END_STRUCT;
      Identification : Struct   // pag 2
         carriage_id_req : Bool;   // Sup->PLC
         new_carriage_id : Bool;   // PLC->Sup
         id_req : Bool;   // Sup->PLC
         id_running : Bool;   // PLC->Sup
         id_ok : Bool;   // PLC->Sup
         teach_req : Bool;   // Sup->PLC
         system_ok : Bool;   // PLC->Sup (parte de id_ok)
         pa_check_req : Bool;   // Sup->PLC
         tcg_req : Bool;   // Sup->PLC
      END_STRUCT;
      Teaching : Struct   // pag 3
         teach_ready : Bool;   // PLC->Sup
         teach_running : Bool;   // Sup->PLC
         teach_state : Bool;   // Sup->PLC
         jump_start_us : Bool;   // PLC->Sup
      END_STRUCT;
      StartUs : Struct   // pag 4
         start_us_ready : Bool;   // PLC->Sup
         start_us_running : Bool;   // Sup->PLC
         start_us_state : Bool;   // Sup->PLC
      END_STRUCT;
      PACheck : Struct   // pag 5
         pa_check_ready : Bool;   // PLC->Sup
         elem_running : Bool;   // Sup->PLC
         elem_state : Bool;   // Sup->PLC
         bal_running : Bool;   // Sup->PLC
         bal_state : Bool;   // Sup->PLC
      END_STRUCT;
      Gain : Struct
         gain_ready : Bool;
         gain_running : Bool;
         gain_state : Bool;
      END_STRUCT;
      TCG_Check : Struct
         tcg_ready : Bool;
         tcg_running : Bool;
         tcg_next_step : Bool;
         jump_acq_ref : Bool;
         jump_tcg_adj : Bool;
      END_STRUCT;
      TCG_Adjust : Struct
         tcg_ready : Bool;
         jump_ref_acq : Bool;
      END_STRUCT;
      RefScan_Acq : Struct
         scan_ref_ready : Bool;
         scan_ref_running : Bool;
      END_STRUCT;
      InspScan : Struct
         scan_insp_ready : Bool;
         scan_insp_running : Bool;
         scan_insp_state : Bool;
         jump_ref_insp : Bool;
      END_STRUCT;
      RefScan_Verif : Struct
         scan_ref_ready : Bool;
         scan_ref_running : Bool;
         jump_start : Bool;
      END_STRUCT;
      Marking : Struct
         mark_req : Bool;
         mark_running : Bool;
         mark_state : Bool;
         jump_start : Bool;
         point_coordinates : Struct
            x : Real;
            y : Real;
            z : Real;
            "a" : Real;
            "b" : Real;
            c : Real;
         END_STRUCT;
      END_STRUCT;
   END_VAR
BEGIN
END_DATA_BLOCK

// folder: System blocks/Program resources

DATA_BLOCK "IEC_Timer_0_DB"   // DB24
{ S7_Optimized_Access := 'TRUE' }
AUTHOR : Simatic
FAMILY : IEC
NAME : IEC_TMR
VERSION : 1.0
// stored: InstanceOfName IEC_TIMER
"IEC_TIMER"
BEGIN
END_DATA_BLOCK

DATA_BLOCK "IEC_Timer_0_DB_1"   // DB25
{ S7_Optimized_Access := 'TRUE' }
AUTHOR : Simatic
FAMILY : IEC
NAME : IEC_TMR
VERSION : 1.0
// stored: InstanceOfName IEC_TIMER
"IEC_TIMER"
BEGIN
END_DATA_BLOCK

DATA_BLOCK "IEC_Timer_0_DB_2"   // DB26
{ S7_Optimized_Access := 'TRUE' }
AUTHOR : Simatic
FAMILY : IEC
NAME : IEC_TMR
VERSION : 1.0
// stored: InstanceOfName IEC_TIMER
"IEC_TIMER"
BEGIN
END_DATA_BLOCK

DATA_BLOCK "IEC_Timer_0_DB_3"   // DB29
{ S7_Optimized_Access := 'TRUE' }
AUTHOR : Simatic
FAMILY : IEC
NAME : IEC_TMR
VERSION : 1.0
// stored: InstanceOfName IEC_TIMER
"IEC_TIMER"
BEGIN
END_DATA_BLOCK

DATA_BLOCK "IEC_Timer_0_DB_4"   // DB30
{ S7_Optimized_Access := 'TRUE' }
AUTHOR : Simatic
FAMILY : IEC
NAME : IEC_TMR
VERSION : 1.0
// stored: InstanceOfName IEC_TIMER
"IEC_TIMER"
BEGIN
END_DATA_BLOCK

DATA_BLOCK "IEC_Timer_0_DB_5"   // DB31
{ S7_Optimized_Access := 'TRUE' }
AUTHOR : Simatic
FAMILY : IEC
NAME : IEC_TMR
VERSION : 1.0
// stored: InstanceOfName IEC_TIMER
"IEC_TIMER"
BEGIN
END_DATA_BLOCK

// folder: (top level)

ORGANIZATION_BLOCK "Startup"   // OB100, LAD, Startup
TITLE = "Complete Restart"
{ S7_Optimized_Access := 'TRUE' }
VERSION : 0.1
   VAR_INPUT
      LostRetentive : Bool;   // True if retentive data are lost
      LostRTC : Bool;   // True if date and time are lost
   END_VAR
BEGIN

REGION Network 1 (SCL): // ====================== READ (%I) ======================
   // // —— Enlaza estos símbolos a tus %I en el árbol de dispositivos ——
   //   // EStop_DI, SafeDoor_DI, AirPressure_DI, WaterInsp_DI, WaterTank_DI, RobotReady_DI, ...
   "$MOVE_ENABLE" := TRUE;
END_REGION
END_ORGANIZATION_BLOCK

// folder: 10. System

FUNCTION_BLOCK "SeqManager"   // FB20, LAD
{ S7_Optimized_Access := 'TRUE' }
VERSION : 0.1
   VAR_INPUT
      systemArmed : Bool;
      autoBusy : Bool;
      servBusy : Bool;
      modeRequest : UInt;
      modeReqSeq : UInt;
   END_VAR
   VAR_OUTPUT
      modeEffective : UInt;
      startAutoExt : Bool;
      enterCellCase1 : Bool;
      enterCellCase2 : Bool;
   END_VAR
   VAR
      lastSeq : UInt;
      safeAllOk : Bool;
      acceptSrv : Bool;
      acceptAuto : Bool;
      firstScan : Bool := true;
   END_VAR
BEGIN

REGION Network 1 (SCL)
   // ----------------- 0) Inicialización por scan -----------------
   "PlcStatus".exec.accepted := FALSE; // pulso hacia la HMI
   "PlcStatus".exec.done := FALSE;    // pulso hacia la HMI

   // Clave: forzamos a FALSE por defecto para que al conceder se produzca pulso
   #startAutoExt := FALSE;
   #enterCellCase2 := FALSE;
   #enterCellCase1 := FALSE;

   // ----------------- 1) Inicialización primera pasada -----------------
   IF  #firstScan THEN
       #firstScan := FALSE;
       #lastSeq := #modeReqSeq;     // ignorar residuos SOLO al arrancar
   END_IF;

   #safeAllOk := #systemArmed;

   // Condición global de seguridad (quedar por ajustar)
   #safeAllOk := #systemArmed;


   IF #modeRequest = 3 THEN
       //#startAutoExt := TRUE;
       #lastSeq := #lastSeq + 1;
       // 5) Handshake a la HMI con el MISMO seq que se recibió
   END_IF;